HMI tags "VAT_PN_PB"
   "PN_PB\PTMUX_P_TLN17_32" : UInt, internal
   "PN_PB\PTMUX_P_TLN1_16" : UInt, internal
   "PN_PB\PTMUX_P_TLN129_144" : UInt, internal
   "PN_PB\DB_PN" : UInt, internal
   "PN_PB\PTMUX_P_TLN177_192" : UInt, internal
   "PN_PB\PTMUX_F_TLN241_256" : UInt, internal
   "PN_PB\IO_Sys_ID" : Int, internal
   "PN_PB\PTMUX_P_TLN225_240" : UInt, internal
   "PN_PB\PTMUX_P_TLN241_256" : UInt, internal
   "PN_PB\PTMUX_P_TLN193_208" : UInt, internal
   "PN_PB\PTMUX_F_TLN1_16" : UInt, internal
   "PN_PB\PTMUX_P_TLN209_224" : UInt, internal
   "PN_PB\PTMUX_F_TLN49_64" : UInt, internal
   "PN_PB\PTMUX_P_TLN113_128" : UInt, internal
   "PN_PB\PTMUX_F_TLN177_192" : UInt, internal
   "PN_PB\PTMUX_P_TLN49_64" : UInt, internal
   "PN_PB\PTMUX_F_TLN97_112" : UInt, internal
   "PN_PB\DB_PB" : UInt, internal
   "PN_PB\PTMUX_F_TLN81_96" : UInt, internal
   "PN_PB\PTMUX_F_TLN145_160" : UInt, internal
   "PN_PB\Diag_Art" : Int, internal
   "PN_PB\PTMUX_F_TLN113_128" : UInt, internal
   "PN_PB\PTMUX_P_TLN97_112" : UInt, internal
   "PN_PB\Teiln_Nr_Anz." : Int, internal
   "PN_PB\PTMUX_P_TLN33_48" : UInt, internal
   "PN_PB\PTMUX_F_TLN161_176" : UInt, internal
   "PN_PB\PTMUX_F_TLN193_208" : UInt, internal
   "PN_PB\PTMUX_P_TLN81_96" : UInt, internal
   "PN_PB\PTMUX_P_TLN65_80" : UInt, internal
   "PN_PB\PTMUX_F_TLN225_240" : UInt, internal
   "PN_PB\PTMUX_F_TLN17_32" : UInt, internal
   "PN_PB\PTMUX_F_TLN65_80" : UInt, internal
   "PN_PB\PTMUX_F_TLN209_224" : UInt, internal
   "PN_PB\PTMUX_F_TLN33_48" : UInt, internal
   "PN_PB\PTMUX_P_TLN145_160" : UInt, internal
   "PN_PB\PTMUX_P_TLN161_176" : UInt, internal
   "PN_PB\Teiln_Nr_Bez" : WString[20], internal
   "PN_PB\Teiln_Nr_Typ" : WString[12], internal
   "PN_PB\Teiln_Nr_Ort" : WString[12], internal
   "PN_PB\PTMUX_F_TLN129_144" : UInt, internal

HMI tags "VAT_SYSTEM_PN"
   "PN_PB\PN\TLN_P_161_176" : Word AT %DB0.DBW230, 100 ms
   "PN_PB\PN\TLN_F_241_256" : Word AT %DB0.DBW368, 100 ms
   "PN_PB\PN\TLN_P_33_48" : Word AT %DB0.DBW214, 100 ms
   "PN_PB\PN\TLN_F_49_64" : Word AT %DB0.DBW344, 100 ms
   "PN_PB\PN\TLN_F_81_96" : Word AT %DB0.DBW348, 100 ms
   "PN_PB\PN\TLN_P_225_240" : Word AT %DB0.DBW238, 100 ms
   "PN_PB\PN\TLN_P_177_192" : Word AT %DB0.DBW232, 100 ms
   "PN_PB\PN\TLN_F_17_32" : Word AT %DB0.DBW340, 100 ms
   "PN_PB\PN\TLN_F_225_240" : Word AT %DB0.DBW366, 100 ms
   "PN_PB\PN\TLN_F_33_48" : Word AT %DB0.DBW342, 100 ms
   "PN_PB\PN\TLN_P_97_112" : Word AT %DB0.DBW222, 100 ms
   "PN_PB\PN\TLN_P_129_144" : Word AT %DB0.DBW226, 100 ms
   "PN_PB\PN\Diag_Slave_Nr" : Int, internal
   "PN_PB\PN\TLN_F_113_128" : Word AT %DB0.DBW352, 100 ms
   "PN_PB\PN\TLN_F_97_112" : Word AT %DB0.DBW350, 100 ms
   "PN_PB\PN\TLN_P_145_160" : Word AT %DB0.DBW228, 100 ms
   "PN_PB\PN\TLN_F_145_160" : Word AT %DB0.DBW356, 100 ms
   "PN_PB\PN\TLN_P_113_128" : Word AT %DB0.DBW224, 100 ms
   "PN_PB\PN\IOSys_ID" : Int AT %DB0.DBW2, 200 ms
   "PN_PB\PN\TLN_F_129_144" : Word AT %DB0.DBW354, 100 ms
   "PN_PB\PN\TLN_F_161_176" : Word AT %DB0.DBW358, 100 ms
   "PN_PB\PN\TLN_F_1_16" : Word AT %DB0.DBW338, 100 ms
   "PN_PB\PN\TLN_P_1_16" : Word AT %DB0.DBW210, 100 ms
   "PN_PB\PN\TLN_P_65_80" : Word AT %DB0.DBW218, 100 ms
   "PN_PB\PN\TLN_F_209_224" : Word AT %DB0.DBW364, 100 ms
   "PN_PB\PN\TLN_F_65_80" : Word AT %DB0.DBW346, 100 ms
   "PN_PB\PN\TLN_P_193_208" : Word AT %DB0.DBW234, 100 ms
   "PN_PB\PN\TLN_P_81_96" : Word AT %DB0.DBW220, 100 ms
   "PN_PB\PN\TLN_P_209_224" : Word AT %DB0.DBW236, 100 ms
   "PN_PB\PN\TLN_P_17_32" : Word AT %DB0.DBW212, 100 ms
   "PN_PB\PN\TLN_P_49_64" : Word AT %DB0.DBW216, 100 ms
   "PN_PB\PN\TLN_P_241_256" : Word AT %DB0.DBW240, 100 ms
   "PN_PB\PN\TLN_F_193_208" : Word AT %DB0.DBW362, 100 ms
   "PN_PB\PN\TLN_F_177_192" : Word AT %DB0.DBW360, 100 ms
   "PN_PB\PN\Teiln_Nr" : Int AT %DB0.DBW4, 1 s
      on ChangeValue: "SDC_PN"()

HMI tags "VAT_SYSTEM_PB"
   "PN_PB\PB\TLN_F_65_80" : Word AT %DB0.DBW234, 100 ms
   "PN_PB\PB\TLN_F_113_128" : Word AT %DB0.DBW240, 100 ms
   "PN_PB\PB\IOSys_ID" : Int AT %DB0.DBW2, 200 ms
   "PN_PB\PB\TLN_P_81_96" : Word AT %DB0.DBW220, 100 ms
   "PN_PB\PB\TLN_F_81_96" : Word AT %DB0.DBW236, 100 ms
   "PN_PB\PB\TLN_F_49_64" : Word AT %DB0.DBW232, 100 ms
   "PN_PB\PB\TLN_P_113_128" : Word AT %DB0.DBW224, 100 ms
   "PN_PB\PB\TLN_F_33_48" : Word AT %DB0.DBW230, 100 ms
   "PN_PB\PB\TLN_P_65_80" : Word AT %DB0.DBW218, 100 ms
   "PN_PB\PB\TLN_P_49_64" : Word AT %DB0.DBW216, 100 ms
   "PN_PB\PB\TLN_F_1_16" : Word AT %DB0.DBW226, 100 ms
   "PN_PB\PB\TLN_P_17_32" : Word AT %DB0.DBW212, 100 ms
   "PN_PB\PB\TLN_P_33_48" : Word AT %DB0.DBW214, 100 ms
   "PN_PB\PB\TLN_P_1_16" : Word AT %DB0.DBW210, 100 ms
   "PN_PB\PB\TLN_F_17_32" : Word AT %DB0.DBW228, 100 ms
   "PN_PB\PB\TLN_F_97_112" : Word AT %DB0.DBW238, 100 ms
   "PN_PB\PB\TLN_P_97_112" : Word AT %DB0.DBW222, 100 ms
   "PN_PB\PB\Teiln_Nr" : Int AT %DB0.DBW4, 200 ms

HMI tags "VAT_SYSTEM_PARAMETER"
   "_intern_Pult_Nr" : Int, internal   // !!! VOR DEM LADEN EINSTELLEN !!!

HMI tags "UserDiag_TagTable"
   "UserDiag_HmiData_actIOSystem" : Int = PLC UserDiag_HmiData.actIOSystem, 1 s
   "UserDiag_HmiData_actDeviceOfScreen" : Int = PLC UserDiag_HmiData.actDeviceOfScreen, 1 s
   "UserDiag_HmiData_ioSlotDiagnosticsLoaded" : Bool = PLC UserDiag_HmiData.ioSlotDiagnosticsLoaded, 1 s
   "UserDiag_HmiData_actScreenDevices" : Int = PLC UserDiag_HmiData.actScreenDevices, 100 ms
   "UserDiag_HmiData_maxScreensDevices" : Int = PLC UserDiag_HmiData.maxScreensDevices, 1 s
   "UserDiag_HmiData_ackWaitTime" : Int = PLC UserDiag_HmiData.ackWaitTime, 1 s
   "UserDiag_HmiData_ackStates" : Bool = PLC UserDiag_HmiData.ackStates, 1 s
   "UserDiag_HmiData_actIOSystemData" : UserDiag_typeActIOSystem = PLC UserDiag_HmiData.actIOSystemData, 1 s
   "UserDiag_HmiData_actDeviceNumber" : UInt = PLC UserDiag_HmiData.actDeviceNumber, 1 s
   "UserDiag_HmiData_actDeviceName" : String[50] = PLC UserDiag_HmiData.actDeviceName, 1 s
   "UserDiag_HmiData_actIPAddress.ADDR" : Array [0..3] of Byte = PLC UserDiag_HmiData.actIPAddress.ADDR, 1 s
   "UserDiag_HmiData_ioSystemError" : Array [0..1] of Bool = PLC UserDiag_HmiData.ioSystemError AT %DB1.DBX0.0, 500 ms
   "UserDiag_HmiData_filterErrorDevices" : Bool = PLC UserDiag_HmiData.filterErrorDevices AT %DB1.DBX0.0, 500 ms
   "UserDiag_HmiData_errorAtLowerScreen" : Bool = PLC UserDiag_HmiData.errorAtLowerScreen, 500 ms
   "UserDiag_HmiData_errorAtUpperScreen" : Bool = PLC UserDiag_HmiData.errorAtUpperScreen AT %DB1.DBW0, 500 ms
   "ioSystem1" : Int AT %DB1.DBW0
   "ioSystem2" : Int AT %DB1.DBW0
   "ioSystem3" : Int AT %DB1.DBW0
   "DB_SDC_FAULTS" : Word = PLC DB101_DB_SDC_FAULTS.SDC_Fault AT %DB101.DBW0, 1 s

HMI tags "DB_SDC_FAULTS"
   "DB101_DB_SDC_FAULTS_SDC_Fault" : Word = PLC DB101_DB_SDC_FAULTS.SDC_Fault AT %DB101.DBW0, 1 s
   "DB101_DB_SDC_FAULTS_Carrier_Fault[15]" : Word = PLC DB101_DB_SDC_FAULTS.Carrier_Fault[15] AT %DB101.DBW30, 1 s
   "DB101_DB_SDC_FAULTS_Carrier_Fault[27]" : Word = PLC DB101_DB_SDC_FAULTS.Carrier_Fault[27] AT %DB101.DBW54, 1 s
   "DB101_DB_SDC_FAULTS_Carrier_Fault[31]" : Word = PLC DB101_DB_SDC_FAULTS.Carrier_Fault[31] AT %DB101.DBW62, 1 s
   "DB101_DB_SDC_FAULTS_Carrier_Fault[40]" : Word = PLC DB101_DB_SDC_FAULTS.Carrier_Fault[40] AT %DB101.DBW80, 1 s

HMI tags "DB_HMI_FAULTS"
   "DB302_HMI_Faults_SDC_Faults_0" : Int = PLC DB302_HMI_Faults.SDC_Faults_0, 1 s
   "DB302_HMI_Faults_SDC_Faults_1" : Int = PLC DB302_HMI_Faults.SDC_Faults_1, 1 s
   "DB302_HMI_Faults_SDC_Faults_2" : Int = PLC DB302_HMI_Faults.SDC_Faults_2, 1 s
   "DB302_HMI_Faults_SDC_Faults_3" : Int = PLC DB302_HMI_Faults.SDC_Faults_3, 1 s

HMI tags "EMS"
   "EMS" : UDT_System = PLC EMS AT %DB1.DBW0, 1 s

HMI tags "DeviceStates_Condition"
   "DB16_EMS_Status_EMS_DeviceStates.DeviceStates_Condition_HMI[2]" : Int = PLC DB16_EMS_Status.EMS_DeviceStates.DeviceStates_Condition_HMI[2], 1 s
   "DB16_EMS_Status_EMS_DeviceStates.DeviceStates_Condition_HMI[3]" : Int = PLC DB16_EMS_Status.EMS_DeviceStates.DeviceStates_Condition_HMI[3], 1 s
   "DB16_EMS_Status_EMS_DeviceStates.DeviceStates_Condition_HMI[4]" : Int = PLC DB16_EMS_Status.EMS_DeviceStates.DeviceStates_Condition_HMI[4], 1 s
   "DB16_EMS_Status_EMS_DeviceStates.DeviceStates_Condition_HMI[5]" : Int = PLC DB16_EMS_Status.EMS_DeviceStates.DeviceStates_Condition_HMI[5], 1 s
   "DB16_EMS_Status_EMS_DeviceStates.DeviceStates_Condition_HMI[6]" : Int = PLC DB16_EMS_Status.EMS_DeviceStates.DeviceStates_Condition_HMI[6], 1 s
   "DB16_EMS_Status_EMS_DeviceStates.DeviceStates_Condition_HMI[7]" : Int = PLC DB16_EMS_Status.EMS_DeviceStates.DeviceStates_Condition_HMI[7], 1 s
   "DB16_EMS_Status_EMS_DeviceStates.DeviceStates_Condition_HMI[8]" : Int = PLC DB16_EMS_Status.EMS_DeviceStates.DeviceStates_Condition_HMI[8], 1 s
   "DB16_EMS_Status_EMS_DeviceStates.DeviceStates_Condition_HMI[9]" : Int = PLC DB16_EMS_Status.EMS_DeviceStates.DeviceStates_Condition_HMI[9], 1 s
   "DB16_EMS_Status_EMS_DeviceStates.DeviceStates_Condition_HMI[10]" : Int = PLC DB16_EMS_Status.EMS_DeviceStates.DeviceStates_Condition_HMI[10], 1 s
   "DB16_EMS_Status_EMS_DeviceStates.DeviceStates_Condition_HMI[11]" : Int = PLC DB16_EMS_Status.EMS_DeviceStates.DeviceStates_Condition_HMI[11], 1 s
   "DB16_EMS_Status_EMS_DeviceStates.DeviceStates_Condition_HMI[12]" : Int = PLC DB16_EMS_Status.EMS_DeviceStates.DeviceStates_Condition_HMI[12], 1 s
   "DB16_EMS_Status_EMS_DeviceStates.DeviceStates_Condition_HMI[13]" : Int = PLC DB16_EMS_Status.EMS_DeviceStates.DeviceStates_Condition_HMI[13], 1 s
   "DB16_EMS_Status_EMS_DeviceStates.DeviceStates_Condition_HMI[14]" : Int = PLC DB16_EMS_Status.EMS_DeviceStates.DeviceStates_Condition_HMI[14], 1 s
   "DB16_EMS_Status_EMS_DeviceStates.DeviceStates_Condition_HMI[15]" : Int = PLC DB16_EMS_Status.EMS_DeviceStates.DeviceStates_Condition_HMI[15], 1 s
   "DB16_EMS_Status_EMS_DeviceStates.DeviceStates_Condition_HMI[16]" : Int = PLC DB16_EMS_Status.EMS_DeviceStates.DeviceStates_Condition_HMI[16], 1 s
   "DB16_EMS_Status_EMS_DeviceStates.DeviceStates_Condition_HMI[17]" : Int = PLC DB16_EMS_Status.EMS_DeviceStates.DeviceStates_Condition_HMI[17], 1 s
   "DB16_EMS_Status_EMS_DeviceStates.DeviceStates_Condition_HMI[18]" : Int = PLC DB16_EMS_Status.EMS_DeviceStates.DeviceStates_Condition_HMI[18], 1 s
   "DB16_EMS_Status_EMS_DeviceStates.DeviceStates_Condition_HMI[19]" : Int = PLC DB16_EMS_Status.EMS_DeviceStates.DeviceStates_Condition_HMI[19], 1 s
   "DB16_EMS_Status_EMS_DeviceStates.DeviceStates_Condition_HMI[20]" : Int = PLC DB16_EMS_Status.EMS_DeviceStates.DeviceStates_Condition_HMI[20], 1 s
   "DB16_EMS_Status_EMS_DeviceStates.DeviceStates_Condition_HMI[21]" : Int = PLC DB16_EMS_Status.EMS_DeviceStates.DeviceStates_Condition_HMI[21], 1 s
   "DB16_EMS_Status_EMS_DeviceStates.DeviceStates_Condition_HMI[22]" : Int = PLC DB16_EMS_Status.EMS_DeviceStates.DeviceStates_Condition_HMI[22], 1 s
   "DB16_EMS_Status_EMS_DeviceStates.DeviceStates_Condition_HMI[23]" : Int = PLC DB16_EMS_Status.EMS_DeviceStates.DeviceStates_Condition_HMI[23], 1 s
   "DB16_EMS_Status_EMS_DeviceStates.DeviceStates_Condition_HMI[24]" : Int = PLC DB16_EMS_Status.EMS_DeviceStates.DeviceStates_Condition_HMI[24], 1 s
   "DB16_EMS_Status_EMS_DeviceStates.DeviceStates_Condition_HMI[25]" : Int = PLC DB16_EMS_Status.EMS_DeviceStates.DeviceStates_Condition_HMI[25], 1 s
   "DB16_EMS_Status_EMS_DeviceStates.DeviceStates_Condition_HMI[26]" : Int = PLC DB16_EMS_Status.EMS_DeviceStates.DeviceStates_Condition_HMI[26], 1 s
   "DB16_EMS_Status_EMS_DeviceStates.DeviceStates_Condition_HMI[27]" : Int = PLC DB16_EMS_Status.EMS_DeviceStates.DeviceStates_Condition_HMI[27], 1 s
   "DB16_EMS_Status_EMS_DeviceStates.DeviceStates_Condition_HMI[28]" : Int = PLC DB16_EMS_Status.EMS_DeviceStates.DeviceStates_Condition_HMI[28], 1 s
   "DB16_EMS_Status_EMS_DeviceStates.DeviceStates_Condition_HMI[29]" : Int = PLC DB16_EMS_Status.EMS_DeviceStates.DeviceStates_Condition_HMI[29], 1 s
   "DB16_EMS_Status_EMS_DeviceStates.DeviceStates_Condition_HMI[30]" : Int = PLC DB16_EMS_Status.EMS_DeviceStates.DeviceStates_Condition_HMI[30], 1 s
   "DB16_EMS_Status_EMS_DeviceStates.DeviceStates_Condition_HMI[31]" : Int = PLC DB16_EMS_Status.EMS_DeviceStates.DeviceStates_Condition_HMI[31], 1 s
   "DB16_EMS_Status_EMS_DeviceStates.DeviceStates_Condition_HMI[32]" : Int = PLC DB16_EMS_Status.EMS_DeviceStates.DeviceStates_Condition_HMI[32], 1 s
   "DB16_EMS_Status_EMS_DeviceStates.DeviceStates_Condition_HMI[33]" : Int = PLC DB16_EMS_Status.EMS_DeviceStates.DeviceStates_Condition_HMI[33], 1 s
   "DB16_EMS_Status_EMS_DeviceStates.DeviceStates_Condition_HMI[34]" : Int = PLC DB16_EMS_Status.EMS_DeviceStates.DeviceStates_Condition_HMI[34], 1 s
   "DB16_EMS_Status_EMS_DeviceStates.DeviceStates_Condition_HMI[35]" : Int = PLC DB16_EMS_Status.EMS_DeviceStates.DeviceStates_Condition_HMI[35], 1 s
   "DB16_EMS_Status_EMS_DeviceStates.DeviceStates_Condition_HMI[36]" : Int = PLC DB16_EMS_Status.EMS_DeviceStates.DeviceStates_Condition_HMI[36], 1 s
   "DB16_EMS_Status_EMS_DeviceStates.DeviceStates_Condition_HMI[37]" : Int = PLC DB16_EMS_Status.EMS_DeviceStates.DeviceStates_Condition_HMI[37], 1 s
   "DB16_EMS_Status_EMS_DeviceStates.DeviceStates_Condition_HMI[38]" : Int = PLC DB16_EMS_Status.EMS_DeviceStates.DeviceStates_Condition_HMI[38], 1 s
   "DB16_EMS_Status_EMS_DeviceStates.DeviceStates_Condition_HMI[39]" : Int = PLC DB16_EMS_Status.EMS_DeviceStates.DeviceStates_Condition_HMI[39], 1 s
   "DB16_EMS_Status_EMS_DeviceStates.DeviceStates_Condition_HMI[40]" : Int = PLC DB16_EMS_Status.EMS_DeviceStates.DeviceStates_Condition_HMI[40], 1 s
   "DB16_EMS_Status_EMS_DeviceStates.DeviceStates_Condition_HMI[41]" : Int = PLC DB16_EMS_Status.EMS_DeviceStates.DeviceStates_Condition_HMI[41], 1 s
   "DB16_EMS_Status_EMS_DeviceStates.DeviceStates_Condition_HMI[42]" : Int = PLC DB16_EMS_Status.EMS_DeviceStates.DeviceStates_Condition_HMI[42], 1 s
   "DB16_EMS_Status_EMS_DeviceStates.DeviceStates_Condition_HMI[43]" : Int = PLC DB16_EMS_Status.EMS_DeviceStates.DeviceStates_Condition_HMI[43], 1 s
   "DB16_EMS_Status_EMS_DeviceStates.DeviceStates_Condition_HMI[44]" : Int = PLC DB16_EMS_Status.EMS_DeviceStates.DeviceStates_Condition_HMI[44], 1 s
   "DB16_EMS_Status_EMS_DeviceStates.DeviceStates_Condition_HMI[45]" : Int = PLC DB16_EMS_Status.EMS_DeviceStates.DeviceStates_Condition_HMI[45], 1 s
   "DB16_EMS_Status_EMS_DeviceStates.DeviceStates_Condition_HMI[46]" : Int = PLC DB16_EMS_Status.EMS_DeviceStates.DeviceStates_Condition_HMI[46], 1 s
   "DB16_EMS_Status_EMS_DeviceStates.DeviceStates_Condition_HMI[47]" : Int = PLC DB16_EMS_Status.EMS_DeviceStates.DeviceStates_Condition_HMI[47], 1 s
   "DB16_EMS_Status_EMS_DeviceStates.DeviceStates_Condition_HMI[48]" : Int = PLC DB16_EMS_Status.EMS_DeviceStates.DeviceStates_Condition_HMI[48], 1 s
   "DB16_EMS_Status_EMS_DeviceStates.DeviceStates_Condition_HMI[49]" : Int = PLC DB16_EMS_Status.EMS_DeviceStates.DeviceStates_Condition_HMI[49], 1 s
   "DB16_EMS_Status_EMS_DeviceStates.DeviceStates_Condition_HMI[50]" : Int = PLC DB16_EMS_Status.EMS_DeviceStates.DeviceStates_Condition_HMI[50], 1 s
   "DB16_EMS_Status_EMS_DeviceStates.DeviceStates_Condition_HMI[51]" : Int = PLC DB16_EMS_Status.EMS_DeviceStates.DeviceStates_Condition_HMI[51], 1 s
   "DB16_EMS_Status_EMS_DeviceStates.DeviceStates_Condition_HMI[52]" : Int = PLC DB16_EMS_Status.EMS_DeviceStates.DeviceStates_Condition_HMI[52], 1 s
   "DB16_EMS_Status_EMS_DeviceStates.DeviceStates_Condition_HMI[53]" : Int = PLC DB16_EMS_Status.EMS_DeviceStates.DeviceStates_Condition_HMI[53], 1 s
   "DB16_EMS_Status_EMS_DeviceStates.DeviceStates_Condition_HMI[54]" : Int = PLC DB16_EMS_Status.EMS_DeviceStates.DeviceStates_Condition_HMI[54], 1 s
   "DB16_EMS_Status_EMS_DeviceStates.DeviceStates_Condition_HMI[55]" : Int = PLC DB16_EMS_Status.EMS_DeviceStates.DeviceStates_Condition_HMI[55], 1 s
   "DB16_EMS_Status_EMS_DeviceStates.DeviceStates_Condition_HMI[56]" : Int = PLC DB16_EMS_Status.EMS_DeviceStates.DeviceStates_Condition_HMI[56], 1 s
   "DB16_EMS_Status_EMS_DeviceStates.DeviceStates_Condition_HMI[57]" : Int = PLC DB16_EMS_Status.EMS_DeviceStates.DeviceStates_Condition_HMI[57], 1 s
   "DB16_EMS_Status_EMS_DeviceStates.DeviceStates_Condition_HMI[58]" : Int = PLC DB16_EMS_Status.EMS_DeviceStates.DeviceStates_Condition_HMI[58], 1 s
   "DB16_EMS_Status_EMS_DeviceStates.DeviceStates_Condition_HMI[59]" : Int = PLC DB16_EMS_Status.EMS_DeviceStates.DeviceStates_Condition_HMI[59], 1 s
   "DB16_EMS_Status_EMS_DeviceStates.DeviceStates_Condition_HMI[60]" : Int = PLC DB16_EMS_Status.EMS_DeviceStates.DeviceStates_Condition_HMI[60], 1 s
   "DB16_EMS_Status_EMS_DeviceStates.DeviceStates_Condition_HMI[61]" : Int = PLC DB16_EMS_Status.EMS_DeviceStates.DeviceStates_Condition_HMI[61], 1 s
   "DB16_EMS_Status_EMS_DeviceStates.DeviceStates_Condition_HMI[62]" : Int = PLC DB16_EMS_Status.EMS_DeviceStates.DeviceStates_Condition_HMI[62], 1 s
   "DB16_EMS_Status_EMS_DeviceStates.DeviceStates_Condition_HMI[63]" : Int = PLC DB16_EMS_Status.EMS_DeviceStates.DeviceStates_Condition_HMI[63], 1 s
   "DB16_EMS_Status_EMS_DeviceStates.DeviceStates_Condition_HMI[64]" : Int = PLC DB16_EMS_Status.EMS_DeviceStates.DeviceStates_Condition_HMI[64], 1 s
   "DB16_EMS_Status_EMS_DeviceStates.DeviceStates_Condition_HMI[65]" : Int = PLC DB16_EMS_Status.EMS_DeviceStates.DeviceStates_Condition_HMI[65], 1 s
   "DB16_EMS_Status_EMS_DeviceStates.DeviceStates_Condition_HMI[66]" : Int = PLC DB16_EMS_Status.EMS_DeviceStates.DeviceStates_Condition_HMI[66], 1 s
   "DB16_EMS_Status_EMS_DeviceStates.DeviceStates_Condition_HMI[67]" : Int = PLC DB16_EMS_Status.EMS_DeviceStates.DeviceStates_Condition_HMI[67], 1 s
   "DB16_EMS_Status_EMS_DeviceStates.DeviceStates_Condition_HMI[68]" : Int = PLC DB16_EMS_Status.EMS_DeviceStates.DeviceStates_Condition_HMI[68], 1 s
   "DB16_EMS_Status_EMS_DeviceStates.DeviceStates_Condition_HMI[69]" : Int = PLC DB16_EMS_Status.EMS_DeviceStates.DeviceStates_Condition_HMI[69], 1 s
   "DB16_EMS_Status_EMS_DeviceStates.DeviceStates_Condition_HMI[70]" : Int = PLC DB16_EMS_Status.EMS_DeviceStates.DeviceStates_Condition_HMI[70], 1 s
   "DB16_EMS_Status_EMS_DeviceStates.DeviceStates_Condition_HMI[71]" : Int = PLC DB16_EMS_Status.EMS_DeviceStates.DeviceStates_Condition_HMI[71], 1 s
   "DB16_EMS_Status_EMS_DeviceStates.DeviceStates_Condition_HMI[72]" : Int = PLC DB16_EMS_Status.EMS_DeviceStates.DeviceStates_Condition_HMI[72], 1 s
   "DB16_EMS_Status_EMS_DeviceStates.DeviceStates_Condition_HMI[73]" : Int = PLC DB16_EMS_Status.EMS_DeviceStates.DeviceStates_Condition_HMI[73], 1 s
   "DB16_EMS_Status_EMS_DeviceStates.DeviceStates_Condition_HMI[74]" : Int = PLC DB16_EMS_Status.EMS_DeviceStates.DeviceStates_Condition_HMI[74], 1 s
   "DB16_EMS_Status_EMS_DeviceStates.DeviceStates_Condition_HMI[75]" : Int = PLC DB16_EMS_Status.EMS_DeviceStates.DeviceStates_Condition_HMI[75], 1 s
   "DB16_EMS_Status_EMS_DeviceStates.DeviceStates_Condition_HMI[76]" : Int = PLC DB16_EMS_Status.EMS_DeviceStates.DeviceStates_Condition_HMI[76], 1 s
   "DB16_EMS_Status_EMS_DeviceStates.DeviceStates_Condition_HMI[77]" : Int = PLC DB16_EMS_Status.EMS_DeviceStates.DeviceStates_Condition_HMI[77], 1 s
   "DB16_EMS_Status_EMS_DeviceStates.DeviceStates_Condition_HMI[78]" : Int = PLC DB16_EMS_Status.EMS_DeviceStates.DeviceStates_Condition_HMI[78], 1 s
   "DB16_EMS_Status_EMS_DeviceStates.DeviceStates_Condition_HMI[79]" : Int = PLC DB16_EMS_Status.EMS_DeviceStates.DeviceStates_Condition_HMI[79], 1 s
   "DB16_EMS_Status_EMS_DeviceStates.DeviceStates_Condition_HMI[80]" : Int = PLC DB16_EMS_Status.EMS_DeviceStates.DeviceStates_Condition_HMI[80], 1 s
   "DB16_EMS_Status_EMS_DeviceStates.DeviceStates_Condition_HMI[81]" : Int = PLC DB16_EMS_Status.EMS_DeviceStates.DeviceStates_Condition_HMI[81], 1 s
   "DB16_EMS_Status_EMS_DeviceStates.DeviceStates_Condition_HMI[82]" : Int = PLC DB16_EMS_Status.EMS_DeviceStates.DeviceStates_Condition_HMI[82], 1 s
   "DB16_EMS_Status_EMS_DeviceStates.DeviceStates_Condition_HMI[1]" : Int = PLC DB16_EMS_Status.EMS_DeviceStates.DeviceStates_Condition_HMI[1], 1 s
   "DB16_EMS_Status_EMS_DeviceStates.DeviceStates_Condition_HMI" : Array [0..82] of Int = PLC DB16_EMS_Status.EMS_DeviceStates.DeviceStates_Condition_HMI AT %DB1.DBW0, 1 s

discrete alarms
   1: 'Rockwell PLC Comm Fault', class No Acknowledgement, trigger "DB302_HMI_Faults_SDC_Faults_0" bit 0
   2: 'Wireless Access Point 1 Comm Fault', class No Acknowledgement, trigger "DB302_HMI_Faults_SDC_Faults_0" bit 1
   3: 'Wireless Access Point 2 Comm Fault', class No Acknowledgement, trigger "DB302_HMI_Faults_SDC_Faults_0" bit 2
   5: 'Wireless Access Point 4 Comm Fault', class No Acknowledgement, trigger "DB302_HMI_Faults_SDC_Faults_0" bit 4
   6: 'Wireless Access Point 5 Comm Fault', class No Acknowledgement, trigger "DB302_HMI_Faults_SDC_Faults_0" bit 5
   7: 'Wireless Access Point 6 Comm Fault', class No Acknowledgement, trigger "DB302_HMI_Faults_SDC_Faults_0" bit 6
   8: 'Wireless Access Point 7 Comm Fault', class No Acknowledgement, trigger "DB302_HMI_Faults_SDC_Faults_0" bit 7
   9: 'Wireless Access Point 8 Comm Fault', class No Acknowledgement, trigger "DB302_HMI_Faults_SDC_Faults_0" bit 8
   10: 'Wireless Access Point 9 Comm Fault', class No Acknowledgement, trigger "DB302_HMI_Faults_SDC_Faults_0" bit 9
   11: 'Wireless Access Point 10 Comm Fault', class No Acknowledgement, trigger "DB302_HMI_Faults_SDC_Faults_0" bit 10
   12: 'Wireless Access Point 11 Comm Fault', class No Acknowledgement, trigger "DB302_HMI_Faults_SDC_Faults_0" bit 11
   13: 'Wireless Access Point 12 Comm Fault', class No Acknowledgement, trigger "DB302_HMI_Faults_SDC_Faults_0" bit 12
   14: 'Wireless Access Point 13 Comm Fault', class No Acknowledgement, trigger "DB302_HMI_Faults_SDC_Faults_0" bit 13
   15: 'Wireless Access Point 14 Comm Fault', class No Acknowledgement, trigger "DB302_HMI_Faults_SDC_Faults_0" bit 14
   16: 'Wireless Access Point 15 Comm Fault', class No Acknowledgement, trigger "DB302_HMI_Faults_SDC_Faults_0" bit 15
   17: 'Wireless Access Point 16 Comm Fault', class No Acknowledgement, trigger "DB302_HMI_Faults_SDC_Faults_1" bit 0
   18: 'Wireless Access Point 17 Comm Fault', class No Acknowledgement, trigger "DB302_HMI_Faults_SDC_Faults_1" bit 1
   19: 'Wireless Access Point 18 Comm Fault', class No Acknowledgement, trigger "DB302_HMI_Faults_SDC_Faults_1" bit 2
   20: 'Wireless Access Point 19 Comm Fault', class No Acknowledgement, trigger "DB302_HMI_Faults_SDC_Faults_1" bit 3
   21: 'Spare_Fault_021', class No Acknowledgement, trigger "DB302_HMI_Faults_SDC_Faults_1" bit 4
   22: 'Spare_Fault_022', class No Acknowledgement, trigger "DB302_HMI_Faults_SDC_Faults_1" bit 5
   23: 'Spare_Fault_023', class No Acknowledgement, trigger "DB302_HMI_Faults_SDC_Faults_1" bit 6
   24: 'Spare_Fault_024', class No Acknowledgement, trigger "DB302_HMI_Faults_SDC_Faults_1" bit 7
   25: 'Duplicate Carrier Fault', class No Acknowledgement, trigger "DB302_HMI_Faults_SDC_Faults_1" bit 8
   26: 'Spare_Fault_026', class No Acknowledgement, trigger "DB302_HMI_Faults_SDC_Faults_1" bit 9
   27: 'EMS01 System E-Stop', class No Acknowledgement, trigger "DB302_HMI_Faults_SDC_Faults_1" bit 10
   28: 'Spare_Fault_028', class No Acknowledgement, trigger "DB302_HMI_Faults_SDC_Faults_1" bit 11
   29: 'Spare_Fault_029', class No Acknowledgement, trigger "DB302_HMI_Faults_SDC_Faults_1" bit 12
   30: 'Spare_Fault_030', class No Acknowledgement, trigger "DB302_HMI_Faults_SDC_Faults_1" bit 13
   31: 'Spare_Fault_031', class No Acknowledgement, trigger "DB302_HMI_Faults_SDC_Faults_1" bit 14
   32: 'Spare_Fault_032', class No Acknowledgement, trigger "DB302_HMI_Faults_SDC_Faults_1" bit 15
   33: 'Spare_Fault_033', class No Acknowledgement, trigger "DB302_HMI_Faults_SDC_Faults_2" bit 0
   34: 'Spare_Fault_034', class No Acknowledgement, trigger "DB302_HMI_Faults_SDC_Faults_2" bit 1
   35: 'Spare_Fault_035', class No Acknowledgement, trigger "DB302_HMI_Faults_SDC_Faults_2" bit 2
   36: 'Spare_Fault_036', class No Acknowledgement, trigger "DB302_HMI_Faults_SDC_Faults_2" bit 3
   37: 'Spare_Fault_037', class No Acknowledgement, trigger "DB302_HMI_Faults_SDC_Faults_2" bit 4
   38: 'Spare_Fault_038', class No Acknowledgement, trigger "DB302_HMI_Faults_SDC_Faults_2" bit 5
   39: 'Spare_Fault_039', class No Acknowledgement, trigger "DB302_HMI_Faults_SDC_Faults_2" bit 6
   40: 'Spare_Fault_040', class No Acknowledgement, trigger "DB302_HMI_Faults_SDC_Faults_2" bit 7
   41: 'Spare_Fault_041', class No Acknowledgement, trigger "DB302_HMI_Faults_SDC_Faults_2" bit 8
   42: 'Spare_Fault_042', class No Acknowledgement, trigger "DB302_HMI_Faults_SDC_Faults_2" bit 9
   43: 'Spare_Fault_043', class No Acknowledgement, trigger "DB302_HMI_Faults_SDC_Faults_2" bit 10
   44: 'Spare_Fault_044', class No Acknowledgement, trigger "DB302_HMI_Faults_SDC_Faults_2" bit 11
   45: 'Spare_Fault_045', class No Acknowledgement, trigger "DB302_HMI_Faults_SDC_Faults_2" bit 12
   46: 'Spare_Fault_046', class No Acknowledgement, trigger "DB302_HMI_Faults_SDC_Faults_2" bit 13
   47: 'Spare_Fault_047', class No Acknowledgement, trigger "DB302_HMI_Faults_SDC_Faults_2" bit 14
   48: 'Spare_Fault_048', class No Acknowledgement, trigger "DB302_HMI_Faults_SDC_Faults_2" bit 15
   49: 'Spare_Fault_049', class No Acknowledgement, trigger "DB302_HMI_Faults_SDC_Faults_3" bit 0
   50: 'Spare_Fault_050', class No Acknowledgement, trigger "DB302_HMI_Faults_SDC_Faults_3" bit 1
   51: 'Spare_Fault_051', class No Acknowledgement, trigger "DB302_HMI_Faults_SDC_Faults_3" bit 2
   52: 'Spare_Fault_052', class No Acknowledgement, trigger "DB302_HMI_Faults_SDC_Faults_3" bit 3
   53: 'Spare_Fault_053', class No Acknowledgement, trigger "DB302_HMI_Faults_SDC_Faults_3" bit 4
   54: 'Spare_Fault_054', class No Acknowledgement, trigger "DB302_HMI_Faults_SDC_Faults_3" bit 5
   55: 'Spare_Fault_055', class No Acknowledgement, trigger "DB302_HMI_Faults_SDC_Faults_3" bit 6
   56: 'Spare_Fault_056', class No Acknowledgement, trigger "DB302_HMI_Faults_SDC_Faults_3" bit 7
   57: 'Spare_Fault_057', class No Acknowledgement, trigger "DB302_HMI_Faults_SDC_Faults_3" bit 8
   58: 'Spare_Fault_058', class No Acknowledgement, trigger "DB302_HMI_Faults_SDC_Faults_3" bit 9
   59: 'Spare_Fault_059', class No Acknowledgement, trigger "DB302_HMI_Faults_SDC_Faults_3" bit 10
   60: 'Spare_Fault_060', class No Acknowledgement, trigger "DB302_HMI_Faults_SDC_Faults_3" bit 11
   61: 'Spare_Fault_061', class No Acknowledgement, trigger "DB302_HMI_Faults_SDC_Faults_3" bit 12
   62: 'Spare_Fault_062', class No Acknowledgement, trigger "DB302_HMI_Faults_SDC_Faults_3" bit 13
   63: 'Spare_Fault_063', class No Acknowledgement, trigger "DB302_HMI_Faults_SDC_Faults_3" bit 14
   64: 'Spare_Fault_064', class No Acknowledgement, trigger "DB302_HMI_Faults_SDC_Faults_3" bit 15
   65: 'Carrier 01 Disconnect Open Power Fault DI11.0', class No Acknowledgement, trigger "DB302_HMI_Faults_Carrier1_Faults_0" bit 0
   66: 'Carrier 01 Drive Profinet Comm Fault', class No Acknowledgement, trigger "DB302_HMI_Faults_Carrier1_Faults_0" bit 1
   67: 'Carrier 01 Production Stop Not Reset', class No Acknowledgement, trigger "DB302_HMI_Faults_Carrier1_Faults_0" bit 2
   68: 'Carrier 01 CB02122 Tripped', class No Acknowledgement, trigger "DB302_HMI_Faults_Carrier1_Faults_0" bit 3
   69: 'Carrier 01 CB02123 Tripped', class No Acknowledgement, trigger "DB302_HMI_Faults_Carrier1_Faults_0" bit 4
   70: 'Carrier 01 AUX1 CB Tripped', class No Acknowledgement, trigger "DB302_HMI_Faults_Carrier1_Faults_0" bit 5
   71: 'Carrier 01 AUX2 CB Tripped', class No Acknowledgement, trigger "DB302_HMI_Faults_Carrier1_Faults_0" bit 6
   72: 'Carrier 01 PLC Not Communicating', class No Acknowledgement, trigger "DB302_HMI_Faults_Carrier1_Faults_0" bit 7
   73: 'Carrier 01 Safe Input Card Fault', class No Acknowledgement, trigger "DB302_HMI_Faults_Carrier1_Faults_0" bit 8
   74: 'Carrier 01 Safe Output Card Fault', class No Acknowledgement, trigger "DB302_HMI_Faults_Carrier1_Faults_0" bit 9
   75: 'Carrier 01 Standard Input Card Fault', class No Acknowledgement, trigger "DB302_HMI_Faults_Carrier1_Faults_0" bit 10
   76: 'Carrier 01 Standard Output Card Fault', class No Acknowledgement, trigger "DB302_HMI_Faults_Carrier1_Faults_0" bit 11
   77: 'Carrier 01 Encoder Position Fault', class No Acknowledgement, trigger "DB302_HMI_Faults_Carrier1_Faults_0" bit 12
   78: 'Carrier 01 Encoder Internal Error', class No Acknowledgement, trigger "DB302_HMI_Faults_Carrier1_Faults_0" bit 13
   79: 'Carrier 01 Encoder Comm Fault', class No Acknowledgement, trigger "DB302_HMI_Faults_Carrier1_Faults_0" bit 14
   80: 'Carrier 01 HMI Comm Fault', class No Acknowledgement, trigger "DB302_HMI_Faults_Carrier1_Faults_0" bit 15
   81: 'Carrier 01 Crash Detection Fault', class No Acknowledgement, trigger "DB302_HMI_Faults_Carrier1_Faults_1" bit 0
   82: 'Carrier 01 Carrier Number Invalid', class No Acknowledgement, trigger "DB302_HMI_Faults_Carrier1_Faults_1" bit 1
   83: 'Carrier 01 Drive: PROFINET configuration error', class No Acknowledgement, trigger "DB302_HMI_Faults_Carrier1_Faults_1" bit 2
   84: 'Carrier 01 Drive: Error internal communications', class No Acknowledgement, trigger "DB302_HMI_Faults_Carrier1_Faults_1" bit 3
   85: 'Carrier 01 Drive: Motor overtemperature', class No Acknowledgement, trigger "DB302_HMI_Faults_Carrier1_Faults_1" bit 4
   86: 'Carrier 01 Drive: Motor overcurrent', class No Acknowledgement, trigger "DB302_HMI_Faults_Carrier1_Faults_1" bit 5
   87: 'Carrier 01 Drive: Infeed or power unit not ready', class No Acknowledgement, trigger "DB302_HMI_Faults_Carrier1_Faults_1" bit 6
   88: 'Carrier 01 Drive: Short-circuit/ground fault detected', class No Acknowledgement, trigger "DB302_HMI_Faults_Carrier1_Faults_1" bit 7
   89: 'Carrier 01 Drive: PROFINET Setpoint timeout', class No Acknowledgement, trigger "DB302_HMI_Faults_Carrier1_Faults_1" bit 8
   90: 'Carrier 01 Power unit: Overcurrent', class No Acknowledgement, trigger "DB302_HMI_Faults_Carrier1_Faults_1" bit 9
   91: 'Carrier 01 Power unit: DC link voltage overvoltage', class No Acknowledgement, trigger "DB302_HMI_Faults_Carrier1_Faults_1" bit 10
   92: 'Carrier 01 Power unit: DC link voltage undervoltage', class No Acknowledgement, trigger "DB302_HMI_Faults_Carrier1_Faults_1" bit 11
   93: 'Carrier 01 Power unit: Line phase failure in main circuit', class No Acknowledgement, trigger "DB302_HMI_Faults_Carrier1_Faults_1" bit 12
   94: 'Carrier 01 Power unit: Phase failure motor cable', class No Acknowledgement, trigger "DB302_HMI_Faults_Carrier1_Faults_1" bit 13
   95: 'Carrier 01 Power unit: Ground fault', class No Acknowledgement, trigger "DB302_HMI_Faults_Carrier1_Faults_1" bit 14
   96: 'Spare_Fault_096', class No Acknowledgement, trigger "DB302_HMI_Faults_Carrier1_Faults_1" bit 15
   97: 'Carrier 01 Motion Off Fault', class No Acknowledgement, trigger "DB302_HMI_Faults_Carrier1_Faults_2" bit 0
   98: 'Carrier 01 Motion On Fault', class No Acknowledgement, trigger "DB302_HMI_Faults_Carrier1_Faults_2" bit 1
   99: 'Carrier 01 Spacing Fault', class No Acknowledgement, trigger "DB302_HMI_Faults_Carrier1_Faults_2" bit 2
   100: 'Carrier 01 Duplicate Carrier Number Fault', class No Acknowledgement, trigger "DB302_HMI_Faults_Carrier1_Faults_2" bit 3
   101: 'Spare_Fault_101', class No Acknowledgement, trigger "DB302_HMI_Faults_Carrier1_Faults_2" bit 4
   102: 'Spare_Fault_102', class No Acknowledgement, trigger "DB302_HMI_Faults_Carrier1_Faults_2" bit 5
   103: 'Spare_Fault_103', class No Acknowledgement, trigger "DB302_HMI_Faults_Carrier1_Faults_2" bit 6
   104: 'Spare_Fault_104', class No Acknowledgement, trigger "DB302_HMI_Faults_Carrier1_Faults_2" bit 7
   105: 'Spare_Fault_105', class No Acknowledgement, trigger "DB302_HMI_Faults_Carrier1_Faults_2" bit 8
   106: 'Spare_Fault_106', class No Acknowledgement, trigger "DB302_HMI_Faults_Carrier1_Faults_2" bit 9
   107: 'Spare_Fault_107', class No Acknowledgement, trigger "DB302_HMI_Faults_Carrier1_Faults_2" bit 10
   108: 'Spare_Fault_108', class No Acknowledgement, trigger "DB302_HMI_Faults_Carrier1_Faults_2" bit 11
   109: 'Spare_Fault_109', class No Acknowledgement, trigger "DB302_HMI_Faults_Carrier1_Faults_2" bit 12
   110: 'Spare_Fault_110', class No Acknowledgement, trigger "DB302_HMI_Faults_Carrier1_Faults_2" bit 13
   111: 'Spare_Fault_111', class No Acknowledgement, trigger "DB302_HMI_Faults_Carrier1_Faults_2" bit 14
   112: 'Spare_Fault_112', class No Acknowledgement, trigger "DB302_HMI_Faults_Carrier1_Faults_2" bit 15
   113: 'Spare_Fault_113', class No Acknowledgement, trigger "DB302_HMI_Faults_Carrier1_Faults_3" bit 0
   114: 'Spare_Fault_114', class No Acknowledgement, trigger "DB302_HMI_Faults_Carrier1_Faults_3" bit 1
   115: 'Spare_Fault_115', class No Acknowledgement, trigger "DB302_HMI_Faults_Carrier1_Faults_3" bit 2
   116: 'Spare_Fault_116', class No Acknowledgement, trigger "DB302_HMI_Faults_Carrier1_Faults_3" bit 3
   117: 'Spare_Fault_117', class No Acknowledgement, trigger "DB302_HMI_Faults_Carrier1_Faults_3" bit 4
   118: 'Spare_Fault_118', class No Acknowledgement, trigger "DB302_HMI_Faults_Carrier1_Faults_3" bit 5
   119: 'Spare_Fault_119', class No Acknowledgement, trigger "DB302_HMI_Faults_Carrier1_Faults_3" bit 6
   120: 'Spare_Fault_120', class No Acknowledgement, trigger "DB302_HMI_Faults_Carrier1_Faults_3" bit 7
   121: 'Spare_Fault_121', class No Acknowledgement, trigger "DB302_HMI_Faults_Carrier1_Faults_3" bit 8
   122: 'Spare_Fault_122', class No Acknowledgement, trigger "DB302_HMI_Faults_Carrier1_Faults_3" bit 9
   123: 'Spare_Fault_123', class No Acknowledgement, trigger "DB302_HMI_Faults_Carrier1_Faults_3" bit 10
   124: 'Spare_Fault_124', class No Acknowledgement, trigger "DB302_HMI_Faults_Carrier1_Faults_3" bit 11
   125: 'Spare_Fault_125', class No Acknowledgement, trigger "DB302_HMI_Faults_Carrier1_Faults_3" bit 12
   126: 'Spare_Fault_126', class No Acknowledgement, trigger "DB302_HMI_Faults_Carrier1_Faults_3" bit 13
   127: 'Spare_Fault_127', class No Acknowledgement, trigger "DB302_HMI_Faults_Carrier1_Faults_3" bit 14
   128: 'Spare_Fault_128', class No Acknowledgement, trigger "DB302_HMI_Faults_Carrier1_Faults_3" bit 15
   129: 'Carrier 02 Disconnect Open Power Fault DI11.0', class No Acknowledgement, trigger "DB302_HMI_Faults_Carrier2_Faults_0" bit 0
   130: 'Carrier 02 Drive Profinet Comm Fault', class No Acknowledgement, trigger "DB302_HMI_Faults_Carrier2_Faults_0" bit 1
   131: 'Carrier 02 Production Stop Not Reset', class No Acknowledgement, trigger "DB302_HMI_Faults_Carrier2_Faults_0" bit 2
   132: 'Carrier 02 CB02122 Tripped', class No Acknowledgement, trigger "DB302_HMI_Faults_Carrier2_Faults_0" bit 3
   133: 'Carrier 02 CB02123 Tripped', class No Acknowledgement, trigger "DB302_HMI_Faults_Carrier2_Faults_0" bit 4
   134: 'Carrier 02 AUX1 CB Tripped', class No Acknowledgement, trigger "DB302_HMI_Faults_Carrier2_Faults_0" bit 5
   135: 'Carrier 02 AUX2 CB Tripped', class No Acknowledgement, trigger "DB302_HMI_Faults_Carrier2_Faults_0" bit 6
   136: 'Carrier 02 PLC Not Communicating', class No Acknowledgement, trigger "DB302_HMI_Faults_Carrier2_Faults_0" bit 7
   137: 'Carrier 02 Safe Input Card Fault', class No Acknowledgement, trigger "DB302_HMI_Faults_Carrier2_Faults_0" bit 8
   138: 'Carrier 02 Safe Output Card Fault', class No Acknowledgement, trigger "DB302_HMI_Faults_Carrier2_Faults_0" bit 9
   139: 'Carrier 02 Standard Input Card Fault', class No Acknowledgement, trigger "DB302_HMI_Faults_Carrier2_Faults_0" bit 10
   140: 'Carrier 02 Standard Output Card Fault', class No Acknowledgement, trigger "DB302_HMI_Faults_Carrier2_Faults_0" bit 11
   141: 'Carrier 02 Encoder Position Fault', class No Acknowledgement, trigger "DB302_HMI_Faults_Carrier2_Faults_0" bit 12
   142: 'Carrier 02 Encoder Internal Error', class No Acknowledgement, trigger "DB302_HMI_Faults_Carrier2_Faults_0" bit 13
   143: 'Carrier 02 Encoder Comm Fault', class No Acknowledgement, trigger "DB302_HMI_Faults_Carrier2_Faults_0" bit 14
   144: 'Carrier 02 HMI Comm Fault', class No Acknowledgement, trigger "DB302_HMI_Faults_Carrier2_Faults_0" bit 15
   145: 'Carrier 02 Crash Detection Fault', class No Acknowledgement, trigger "DB302_HMI_Faults_Carrier2_Faults_1" bit 0
   146: 'Carrier 02 Carrier Number Invalid', class No Acknowledgement, trigger "DB302_HMI_Faults_Carrier2_Faults_1" bit 1
   147: 'Carrier 02 Drive: PROFINET configuration error', class No Acknowledgement, trigger "DB302_HMI_Faults_Carrier2_Faults_1" bit 2
   148: 'Carrier 02 Drive: Error internal communications', class No Acknowledgement, trigger "DB302_HMI_Faults_Carrier2_Faults_1" bit 3
   149: 'Carrier 02 Drive: Motor overtemperature', class No Acknowledgement, trigger "DB302_HMI_Faults_Carrier2_Faults_1" bit 4
   150: 'Carrier 02 Drive: Motor overcurrent', class No Acknowledgement, trigger "DB302_HMI_Faults_Carrier2_Faults_1" bit 5
   151: 'Carrier 02 Drive: Infeed or power unit not ready', class No Acknowledgement, trigger "DB302_HMI_Faults_Carrier2_Faults_1" bit 6
   152: 'Carrier 02 Drive: Short-circuit/ground fault detected', class No Acknowledgement, trigger "DB302_HMI_Faults_Carrier2_Faults_1" bit 7
   153: 'Carrier 02 Drive: PROFINET Setpoint timeout', class No Acknowledgement, trigger "DB302_HMI_Faults_Carrier2_Faults_1" bit 8
   154: 'Carrier 02 Power unit: Overcurrent', class No Acknowledgement, trigger "DB302_HMI_Faults_Carrier2_Faults_1" bit 9
   155: 'Carrier 02 Power unit: DC link voltage overvoltage', class No Acknowledgement, trigger "DB302_HMI_Faults_Carrier2_Faults_1" bit 10
   156: 'Carrier 02 Power unit: DC link voltage undervoltage', class No Acknowledgement, trigger "DB302_HMI_Faults_Carrier2_Faults_1" bit 11
   157: 'Carrier 02 Power unit: Line phase failure in main circuit', class No Acknowledgement, trigger "DB302_HMI_Faults_Carrier2_Faults_1" bit 12
   158: 'Carrier 02 Power unit: Phase failure motor cable', class No Acknowledgement, trigger "DB302_HMI_Faults_Carrier2_Faults_1" bit 13
   159: 'Carrier 02 Power unit: Ground fault', class No Acknowledgement, trigger "DB302_HMI_Faults_Carrier2_Faults_1" bit 14
   160: 'Spare_Fault_160', class No Acknowledgement, trigger "DB302_HMI_Faults_Carrier2_Faults_1" bit 15
   161: 'Carrier 02 Motion Off Fault', class No Acknowledgement, trigger "DB302_HMI_Faults_Carrier2_Faults_2" bit 0
   162: 'Carrier 02 Motion On Fault', class No Acknowledgement, trigger "DB302_HMI_Faults_Carrier2_Faults_2" bit 1
   163: 'Carrier 02 Spacing Fault', class No Acknowledgement, trigger "DB302_HMI_Faults_Carrier2_Faults_2" bit 2
   164: 'Carrier 02 Duplicate Carrier Number Fault', class No Acknowledgement, trigger "DB302_HMI_Faults_Carrier2_Faults_2" bit 3
   165: 'Spare_Fault_165', class No Acknowledgement, trigger "DB302_HMI_Faults_Carrier2_Faults_2" bit 4
   166: 'Spare_Fault_166', class No Acknowledgement, trigger "DB302_HMI_Faults_Carrier2_Faults_2" bit 5
   167: 'Spare_Fault_167', class No Acknowledgement, trigger "DB302_HMI_Faults_Carrier2_Faults_2" bit 6
   168: 'Spare_Fault_168', class No Acknowledgement, trigger "DB302_HMI_Faults_Carrier2_Faults_2" bit 7
   169: 'Spare_Fault_169', class No Acknowledgement, trigger "DB302_HMI_Faults_Carrier2_Faults_2" bit 8
   170: 'Spare_Fault_170', class No Acknowledgement, trigger "DB302_HMI_Faults_Carrier2_Faults_2" bit 9
   171: 'Spare_Fault_171', class No Acknowledgement, trigger "DB302_HMI_Faults_Carrier2_Faults_2" bit 10
   172: 'Spare_Fault_172', class No Acknowledgement, trigger "DB302_HMI_Faults_Carrier2_Faults_2" bit 11
   173: 'Spare_Fault_173', class No Acknowledgement, trigger "DB302_HMI_Faults_Carrier2_Faults_2" bit 12
   174: 'Spare_Fault_174', class No Acknowledgement, trigger "DB302_HMI_Faults_Carrier2_Faults_2" bit 13
   175: 'Spare_Fault_175', class No Acknowledgement, trigger "DB302_HMI_Faults_Carrier2_Faults_2" bit 14
   176: 'Spare_Fault_176', class No Acknowledgement, trigger "DB302_HMI_Faults_Carrier2_Faults_2" bit 15
   177: 'Spare_Fault_177', class No Acknowledgement, trigger "DB302_HMI_Faults_Carrier2_Faults_3" bit 0
   178: 'Spare_Fault_178', class No Acknowledgement, trigger "DB302_HMI_Faults_Carrier2_Faults_3" bit 1
   179: 'Spare_Fault_179', class No Acknowledgement, trigger "DB302_HMI_Faults_Carrier2_Faults_3" bit 2
   180: 'Spare_Fault_180', class No Acknowledgement, trigger "DB302_HMI_Faults_Carrier2_Faults_3" bit 3
   181: 'Spare_Fault_181', class No Acknowledgement, trigger "DB302_HMI_Faults_Carrier2_Faults_3" bit 4
   182: 'Spare_Fault_182', class No Acknowledgement, trigger "DB302_HMI_Faults_Carrier2_Faults_3" bit 5
   183: 'Spare_Fault_183', class No Acknowledgement, trigger "DB302_HMI_Faults_Carrier2_Faults_3" bit 6
   184: 'Spare_Fault_184', class No Acknowledgement, trigger "DB302_HMI_Faults_Carrier2_Faults_3" bit 7
   185: 'Spare_Fault_185', class No Acknowledgement, trigger "DB302_HMI_Faults_Carrier2_Faults_3" bit 8
   186: 'Spare_Fault_186', class No Acknowledgement, trigger "DB302_HMI_Faults_Carrier2_Faults_3" bit 9
   187: 'Spare_Fault_187', class No Acknowledgement, trigger "DB302_HMI_Faults_Carrier2_Faults_3" bit 10
   188: 'Spare_Fault_188', class No Acknowledgement, trigger "DB302_HMI_Faults_Carrier2_Faults_3" bit 11
   189: 'Spare_Fault_189', class No Acknowledgement, trigger "DB302_HMI_Faults_Carrier2_Faults_3" bit 12
   190: 'Spare_Fault_190', class No Acknowledgement, trigger "DB302_HMI_Faults_Carrier2_Faults_3" bit 13
   191: 'Spare_Fault_191', class No Acknowledgement, trigger "DB302_HMI_Faults_Carrier2_Faults_3" bit 14
   192: 'Spare_Fault_192', class No Acknowledgement, trigger "DB302_HMI_Faults_Carrier2_Faults_3" bit 15
   193: 'Carrier 03 Disconnect Open Power Fault DI11.0', class No Acknowledgement, trigger "DB302_HMI_Faults_Carrier3_Faults_0" bit 0
   194: 'Carrier 03 Drive Profinet Comm Fault', class No Acknowledgement, trigger "DB302_HMI_Faults_Carrier3_Faults_0" bit 1
   195: 'Carrier 03 Production Stop Not Reset', class No Acknowledgement, trigger "DB302_HMI_Faults_Carrier3_Faults_0" bit 2
   196: 'Carrier 03 CB02122 Tripped', class No Acknowledgement, trigger "DB302_HMI_Faults_Carrier3_Faults_0" bit 3
   197: 'Carrier 03 CB02123 Tripped', class No Acknowledgement, trigger "DB302_HMI_Faults_Carrier3_Faults_0" bit 4
   198: 'Carrier 03 AUX1 CB Tripped', class No Acknowledgement, trigger "DB302_HMI_Faults_Carrier3_Faults_0" bit 5
   199: 'Carrier 03 AUX2 CB Tripped', class No Acknowledgement, trigger "DB302_HMI_Faults_Carrier3_Faults_0" bit 6
   200: 'Carrier 03 PLC Not Communicating', class No Acknowledgement, trigger "DB302_HMI_Faults_Carrier3_Faults_0" bit 7
   201: 'Carrier 03 Safe Input Card Fault', class No Acknowledgement, trigger "DB302_HMI_Faults_Carrier3_Faults_0" bit 8
   202: 'Carrier 03 Safe Output Card Fault', class No Acknowledgement, trigger "DB302_HMI_Faults_Carrier3_Faults_0" bit 9
   203: 'Carrier 03 Standard Input Card Fault', class No Acknowledgement, trigger "DB302_HMI_Faults_Carrier3_Faults_0" bit 10
   204: 'Carrier 03 Standard Output Card Fault', class No Acknowledgement, trigger "DB302_HMI_Faults_Carrier3_Faults_0" bit 11
   205: 'Carrier 03 Encoder Position Fault', class No Acknowledgement, trigger "DB302_HMI_Faults_Carrier3_Faults_0" bit 12
   206: 'Carrier 03 Encoder Internal Error', class No Acknowledgement, trigger "DB302_HMI_Faults_Carrier3_Faults_0" bit 13
   207: 'Carrier 03 Encoder Comm Fault', class No Acknowledgement, trigger "DB302_HMI_Faults_Carrier3_Faults_0" bit 14
   208: 'Carrier 03 HMI Comm Fault', class No Acknowledgement, trigger "DB302_HMI_Faults_Carrier3_Faults_0" bit 15
   209: 'Carrier 03 Crash Detection Fault', class No Acknowledgement, trigger "DB302_HMI_Faults_Carrier3_Faults_1" bit 0
   210: 'Carrier 03 Carrier Number Invalid', class No Acknowledgement, trigger "DB302_HMI_Faults_Carrier3_Faults_1" bit 1
   211: 'Carrier 03 Drive: PROFINET configuration error', class No Acknowledgement, trigger "DB302_HMI_Faults_Carrier3_Faults_1" bit 2
   212: 'Carrier 03 Drive: Error internal communications', class No Acknowledgement, trigger "DB302_HMI_Faults_Carrier3_Faults_1" bit 3
   213: 'Carrier 03 Drive: Motor overtemperature', class No Acknowledgement, trigger "DB302_HMI_Faults_Carrier3_Faults_1" bit 4
   214: 'Carrier 03 Drive: Motor overcurrent', class No Acknowledgement, trigger "DB302_HMI_Faults_Carrier3_Faults_1" bit 5
   215: 'Carrier 03 Drive: Infeed or power unit not ready', class No Acknowledgement, trigger "DB302_HMI_Faults_Carrier3_Faults_1" bit 6
   216: 'Carrier 03 Drive: Short-circuit/ground fault detected', class No Acknowledgement, trigger "DB302_HMI_Faults_Carrier3_Faults_1" bit 7
   217: 'Carrier 03 Drive: PROFINET Setpoint timeout', class No Acknowledgement, trigger "DB302_HMI_Faults_Carrier3_Faults_1" bit 8
   218: 'Carrier 03 Power unit: Overcurrent', class No Acknowledgement, trigger "DB302_HMI_Faults_Carrier3_Faults_1" bit 9
   219: 'Carrier 03 Power unit: DC link voltage overvoltage', class No Acknowledgement, trigger "DB302_HMI_Faults_Carrier3_Faults_1" bit 10
   220: 'Carrier 03 Power unit: DC link voltage undervoltage', class No Acknowledgement, trigger "DB302_HMI_Faults_Carrier3_Faults_1" bit 11
   221: 'Carrier 03 Power unit: Line phase failure in main circuit', class No Acknowledgement, trigger "DB302_HMI_Faults_Carrier3_Faults_1" bit 12
   222: 'Carrier 03 Power unit: Phase failure motor cable', class No Acknowledgement, trigger "DB302_HMI_Faults_Carrier3_Faults_1" bit 13
   223: 'Carrier 03 Power unit: Ground fault', class No Acknowledgement, trigger "DB302_HMI_Faults_Carrier3_Faults_1" bit 14
   224: 'Spare_Fault_224', class No Acknowledgement, trigger "DB302_HMI_Faults_Carrier3_Faults_1" bit 15
   225: 'Carrier 03 Motion Off Fault', class No Acknowledgement, trigger "DB302_HMI_Faults_Carrier3_Faults_2" bit 0
   226: 'Carrier 03 Motion On Fault', class No Acknowledgement, trigger "DB302_HMI_Faults_Carrier3_Faults_2" bit 1
   227: 'Carrier 03 Spacing Fault', class No Acknowledgement, trigger "DB302_HMI_Faults_Carrier3_Faults_2" bit 2
   228: 'Carrier 03 Duplicate Carrier Number Fault', class No Acknowledgement, trigger "DB302_HMI_Faults_Carrier3_Faults_2" bit 3
   229: 'Spare_Fault_229', class No Acknowledgement, trigger "DB302_HMI_Faults_Carrier3_Faults_2" bit 4
   230: 'Spare_Fault_230', class No Acknowledgement, trigger "DB302_HMI_Faults_Carrier3_Faults_2" bit 5
   231: 'Spare_Fault_231', class No Acknowledgement, trigger "DB302_HMI_Faults_Carrier3_Faults_2" bit 6
   232: 'Spare_Fault_232', class No Acknowledgement, trigger "DB302_HMI_Faults_Carrier3_Faults_2" bit 7
   233: 'Spare_Fault_233', class No Acknowledgement, trigger "DB302_HMI_Faults_Carrier3_Faults_2" bit 8
   234: 'Spare_Fault_234', class No Acknowledgement, trigger "DB302_HMI_Faults_Carrier3_Faults_2" bit 9
   235: 'Spare_Fault_235', class No Acknowledgement, trigger "DB302_HMI_Faults_Carrier3_Faults_2" bit 10
   236: 'Spare_Fault_236', class No Acknowledgement, trigger "DB302_HMI_Faults_Carrier3_Faults_2" bit 11
   237: 'Spare_Fault_237', class No Acknowledgement, trigger "DB302_HMI_Faults_Carrier3_Faults_2" bit 12
   238: 'Spare_Fault_238', class No Acknowledgement, trigger "DB302_HMI_Faults_Carrier3_Faults_2" bit 13
   239: 'Spare_Fault_239', class No Acknowledgement, trigger "DB302_HMI_Faults_Carrier3_Faults_2" bit 14
   240: 'Spare_Fault_240', class No Acknowledgement, trigger "DB302_HMI_Faults_Carrier3_Faults_2" bit 15
   241: 'Spare_Fault_241', class No Acknowledgement, trigger "DB302_HMI_Faults_Carrier3_Faults_3" bit 0
   242: 'Spare_Fault_242', class No Acknowledgement, trigger "DB302_HMI_Faults_Carrier3_Faults_3" bit 1
   243: 'Spare_Fault_243', class No Acknowledgement, trigger "DB302_HMI_Faults_Carrier3_Faults_3" bit 2
   244: 'Spare_Fault_244', class No Acknowledgement, trigger "DB302_HMI_Faults_Carrier3_Faults_3" bit 3
   245: 'Spare_Fault_245', class No Acknowledgement, trigger "DB302_HMI_Faults_Carrier3_Faults_3" bit 4
   246: 'Spare_Fault_246', class No Acknowledgement, trigger "DB302_HMI_Faults_Carrier3_Faults_3" bit 5
   247: 'Spare_Fault_247', class No Acknowledgement, trigger "DB302_HMI_Faults_Carrier3_Faults_3" bit 6
   248: 'Spare_Fault_248', class No Acknowledgement, trigger "DB302_HMI_Faults_Carrier3_Faults_3" bit 7
   249: 'Spare_Fault_249', class No Acknowledgement, trigger "DB302_HMI_Faults_Carrier3_Faults_3" bit 8
   250: 'Spare_Fault_250', class No Acknowledgement, trigger "DB302_HMI_Faults_Carrier3_Faults_3" bit 9
   251: 'Spare_Fault_251', class No Acknowledgement, trigger "DB302_HMI_Faults_Carrier3_Faults_3" bit 10
   252: 'Spare_Fault_252', class No Acknowledgement, trigger "DB302_HMI_Faults_Carrier3_Faults_3" bit 11
   253: 'Spare_Fault_253', class No Acknowledgement, trigger "DB302_HMI_Faults_Carrier3_Faults_3" bit 12
   254: 'Spare_Fault_254', class No Acknowledgement, trigger "DB302_HMI_Faults_Carrier3_Faults_3" bit 13
   255: 'Spare_Fault_255', class No Acknowledgement, trigger "DB302_HMI_Faults_Carrier3_Faults_3" bit 14
   256: 'Spare_Fault_256', class No Acknowledgement, trigger "DB302_HMI_Faults_Carrier3_Faults_3" bit 15
   257: 'Carrier 04 Disconnect Open Power Fault DI11.0', class No Acknowledgement, trigger "DB302_HMI_Faults_Carrier4_Faults_0" bit 0
   258: 'Carrier 04 Drive Profinet Comm Fault', class No Acknowledgement, trigger "DB302_HMI_Faults_Carrier4_Faults_0" bit 1
   259: 'Carrier 04 Production Stop Not Reset', class No Acknowledgement, trigger "DB302_HMI_Faults_Carrier4_Faults_0" bit 2
   260: 'Carrier 04 CB02122 Tripped', class No Acknowledgement, trigger "DB302_HMI_Faults_Carrier4_Faults_0" bit 3
   261: 'Carrier 04 CB02123 Tripped', class No Acknowledgement, trigger "DB302_HMI_Faults_Carrier4_Faults_0" bit 4
   262: 'Carrier 04 AUX1 CB Tripped', class No Acknowledgement, trigger "DB302_HMI_Faults_Carrier4_Faults_0" bit 5
   263: 'Carrier 04 AUX2 CB Tripped', class No Acknowledgement, trigger "DB302_HMI_Faults_Carrier4_Faults_0" bit 6
   264: 'Carrier 04 PLC Not Communicating', class No Acknowledgement, trigger "DB302_HMI_Faults_Carrier4_Faults_0" bit 7
   265: 'Carrier 04 Safe Input Card Fault', class No Acknowledgement, trigger "DB302_HMI_Faults_Carrier4_Faults_0" bit 8